// TIA Portal project "Star-Delta Motor Starter with Industrial HMI+Fault Protection" (V20)

(* hardware
DEVICE "S7-1200 station_1"  S7-1200 Station
   slot 0: "Rack_0"  S7-1200 Rack  Rack  V1.0
   slot 1: "PLC_1"  CPU 1214C DC/DC/DC  6ES7 214-1AG40-0XB0  V4.7
DEVICE "HMI_1"  KTP700 Basic PN
   slot 0: "HMI_1"  KTP700 Basic PN  6AV2 123-2GB03-0AX0  17.0.0.0
   slot 1: "HMI_RT_1"  KTP700 Basic PN  6AV2 123-2GB03-0AX0  17.0.0.0
   slot 5: "HMI_1.IE_CP_1"  PROFINET Interface  17.0.0.0
      slot 1: "PROFINET Interface_1"  PROFINET Interface
         slot 1: "Port_1"  Port
*)

// ===== PLC "PLC_1"  CPU 1214C DC/DC/DC =====

VAR_GLOBAL   // PLC tag table "Default tag table"
   "Start_PB" AT %I0.0 : Bool;
   "Stop_PB" AT %I0.1 : Bool;
   "Emergency_Stop" AT %I0.2 : Bool;
   "Thermal_Overload" AT %I0.3 : Bool;
   "Phase_Loss_Sensor" AT %I0.4 : Bool;
   "Reset_PB" AT %I0.5 : Bool;
   "Main_Contactor_K1" AT %Q0.0 : Bool;
   "Star_Contactor_K2" AT %Q0.1 : Bool;
   "Delta_Contactor_K3" AT %Q0.2 : Bool;
   "Alarm_Lamp" AT %M10.3 : Bool;
   "Motor_Run_Latch" AT %M0.0 : Bool;
   "Star_Mode" AT %M0.1 : Bool;
   "Delta_Mode" AT %M0.2 : Bool;
   "Fault_Active" AT %M0.3 : Bool;
   "HMI_Start" AT %M0.4 : Bool;
   "HMI_Stop" AT %M0.5 : Bool;
   "HMI_Reset" AT %M0.6 : Bool;
   "Transition_Done" AT %M0.7 : Bool;
   "Start_Command" AT %M1.0 : Bool;
   "Stop_Command" AT %M1.1 : Bool;
   "Star_Timer_Done" AT %M1.2 : Bool;
   "Star_Lamp" AT %M10.2 : Bool;
   "Delta_Lamp" AT %M10.1 : Bool;
   "Start_Pulse" AT %M1.3 : Bool;
END_VAR

DATA_BLOCK "DB_StarDelta"   // DB1
{ S7_Optimized_Access := 'TRUE' }
VERSION : 0.1
   VAR
      Star_timer_Preset : Time := T#5s;
      Transition_Delay : Time := T#500ms;
      Running_Hours : Real := 0.0;
      Start_Counter : Int := 0;
      Fault_Code : Int := 0;
      Motor_Status : Bool;
      Thermal_Alarm : Bool;
      Phase_Loss_Alarm : Bool;
      Star_Contactor_Fault : Bool;
      Delta_Contactor_Fault : Bool;
   END_VAR
BEGIN
END_DATA_BLOCK

// folder: System blocks/Program resources

DATA_BLOCK "Star_Timer"   // DB2
{ S7_Optimized_Access := 'TRUE' }
AUTHOR : Simatic
FAMILY : IEC
NAME : IEC_TMR
VERSION : 1.0
// stored: InstanceOfName IEC_TIMER
"IEC_TIMER"
BEGIN
END_DATA_BLOCK

DATA_BLOCK "Transition_Timer"   // DB3
{ S7_Optimized_Access := 'TRUE' }
AUTHOR : Simatic
FAMILY : IEC
NAME : IEC_TMR
VERSION : 1.0
// stored: InstanceOfName IEC_TIMER
"IEC_TIMER"
BEGIN
END_DATA_BLOCK

// folder: (top level)

ORGANIZATION_BLOCK "Main"   // OB1, LAD, ProgramCycle
TITLE = "Main Program Sweep (Cycle)"
{ S7_Optimized_Access := 'TRUE' }
VERSION : 0.1
   VAR_INPUT
      Initial_Call : Bool;   // Initial call of this OB
      Remanence : Bool;   // =True, if remanent data are available
   END_VAR
BEGIN

REGION Network 1: Start command
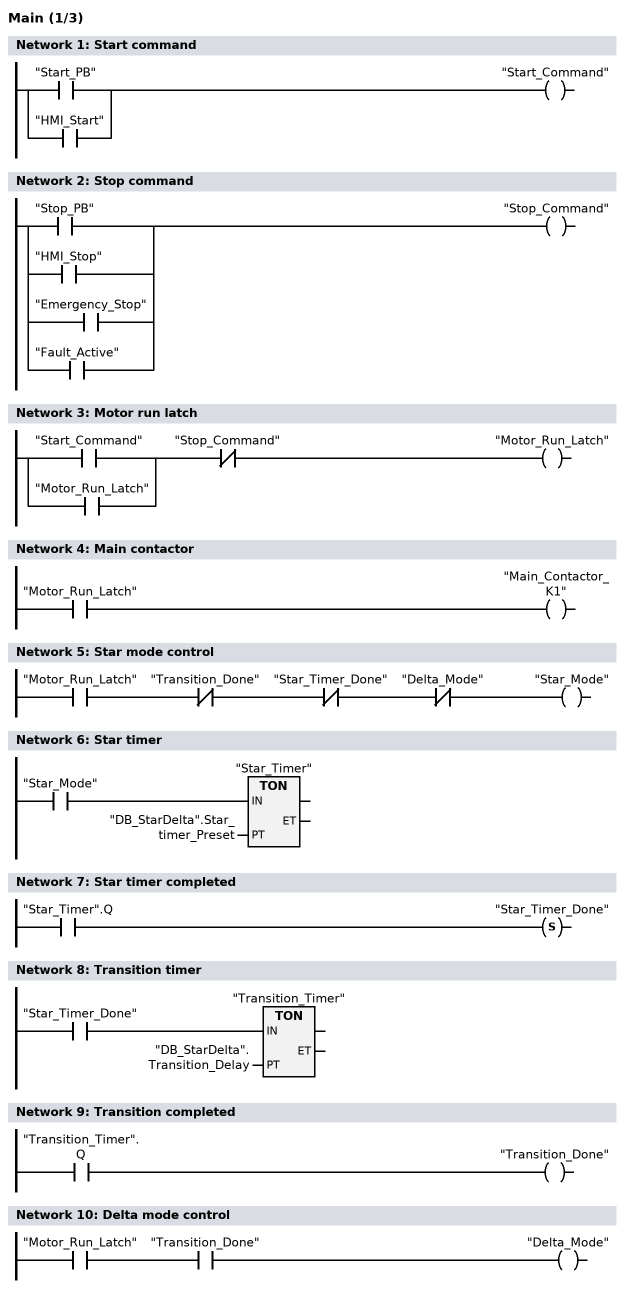
   RUNG wire#powerrail
      Contact( "Start_PB" )
      wire#w1
      Coil( "Start_Command" )
   END_RUNG
   RUNG wire#powerrail
      Contact( "HMI_Start" )
   END_RUNG wire#w1
   // the same network as SCL:
   "Start_Command" := "Start_PB" OR "HMI_Start";
END_REGION

REGION Network 2: Stop command
   RUNG wire#powerrail
      Contact( "Stop_PB" )
      wire#w1
      Coil( "Stop_Command" )
   END_RUNG
   RUNG wire#powerrail
      Contact( "HMI_Stop" )
   END_RUNG wire#w1
   RUNG wire#powerrail
      Contact( "Emergency_Stop" )
   END_RUNG wire#w1
   RUNG wire#powerrail
      Contact( "Fault_Active" )
   END_RUNG wire#w1
   // the same network as SCL:
   "Stop_Command" := "Stop_PB" OR "HMI_Stop" OR "Emergency_Stop" OR "Fault_Active";
END_REGION

REGION Network 3: Motor run latch
   RUNG wire#powerrail
      Contact( "Start_Command" )
      wire#w1
      I_Contact( "Stop_Command" )
      Coil( "Motor_Run_Latch" )
   END_RUNG
   RUNG wire#powerrail
      Contact( "Motor_Run_Latch" )
   END_RUNG wire#w1
   // the same network as SCL:
   "Motor_Run_Latch" := ("Start_Command" OR "Motor_Run_Latch") AND NOT "Stop_Command";
END_REGION

REGION Network 4: Main contactor
   RUNG wire#powerrail
      Contact( "Motor_Run_Latch" )
      Coil( "Main_Contactor_K1" )
   END_RUNG
   // the same network as SCL:
   "Main_Contactor_K1" := "Motor_Run_Latch";
END_REGION

REGION Network 5: Star mode control
   RUNG wire#powerrail
      Contact( "Motor_Run_Latch" )
      I_Contact( "Transition_Done" )
      I_Contact( "Star_Timer_Done" )
      I_Contact( "Delta_Mode" )
      Coil( "Star_Mode" )
   END_RUNG
   // the same network as SCL:
   "Star_Mode" := "Motor_Run_Latch" AND NOT "Transition_Done" AND NOT "Star_Timer_Done" AND NOT "Delta_Mode";
END_REGION

REGION Network 6: Star timer
   "Star_Timer".TON(IN := "Star_Mode", PT := "DB_StarDelta".Star_timer_Preset);
END_REGION

REGION Network 7: Star timer completed
   RUNG wire#powerrail
      Contact( "Star_Timer".Q )
      S_Coil( "Star_Timer_Done" )
   END_RUNG
   // the same network as SCL:
   IF "Star_Timer".Q THEN "Star_Timer_Done" := TRUE; END_IF;
END_REGION

REGION Network 8: Transition timer
   "Transition_Timer".TON(IN := "Star_Timer_Done", PT := "DB_StarDelta".Transition_Delay);
END_REGION

REGION Network 9: Transition completed
   RUNG wire#powerrail
      Contact( "Transition_Timer".Q )
      Coil( "Transition_Done" )
   END_RUNG
   // the same network as SCL:
   "Transition_Done" := "Transition_Timer".Q;
END_REGION

REGION Network 10: Delta mode control
   RUNG wire#powerrail
      Contact( "Motor_Run_Latch" )
      Contact( "Transition_Done" )
      Coil( "Delta_Mode" )
   END_RUNG
   // the same network as SCL:
   "Delta_Mode" := "Motor_Run_Latch" AND "Transition_Done";
END_REGION

REGION Network 11: Delta contactor
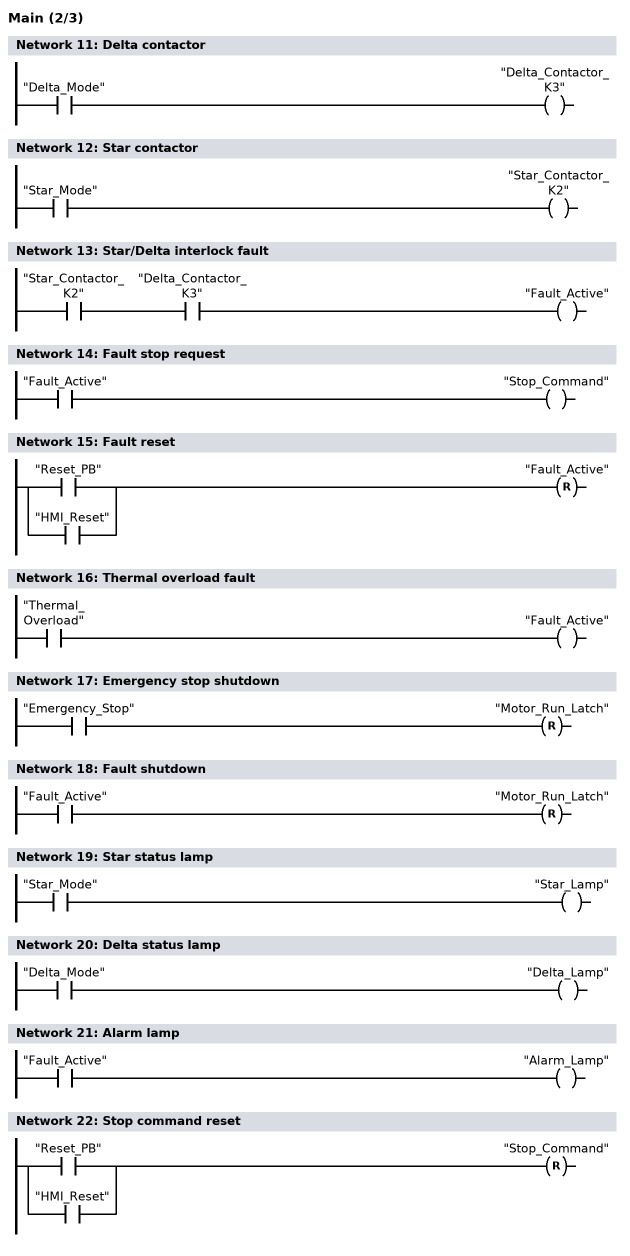
   RUNG wire#powerrail
      Contact( "Delta_Mode" )
      Coil( "Delta_Contactor_K3" )
   END_RUNG
   // the same network as SCL:
   "Delta_Contactor_K3" := "Delta_Mode";
END_REGION

REGION Network 12: Star contactor
   RUNG wire#powerrail
      Contact( "Star_Mode" )
      Coil( "Star_Contactor_K2" )
   END_RUNG
   // the same network as SCL:
   "Star_Contactor_K2" := "Star_Mode";
END_REGION

REGION Network 13: Star/Delta interlock fault
   RUNG wire#powerrail
      Contact( "Star_Contactor_K2" )
      Contact( "Delta_Contactor_K3" )
      Coil( "Fault_Active" )
   END_RUNG
   // the same network as SCL:
   "Fault_Active" := "Star_Contactor_K2" AND "Delta_Contactor_K3";
END_REGION

REGION Network 14: Fault stop request
   RUNG wire#powerrail
      Contact( "Fault_Active" )
      Coil( "Stop_Command" )
   END_RUNG
   // the same network as SCL:
   "Stop_Command" := "Fault_Active";
END_REGION

REGION Network 15: Fault reset
   RUNG wire#powerrail
      Contact( "Reset_PB" )
      wire#w1
      R_Coil( "Fault_Active" )
   END_RUNG
   RUNG wire#powerrail
      Contact( "HMI_Reset" )
   END_RUNG wire#w1
   // the same network as SCL:
   IF "Reset_PB" OR "HMI_Reset" THEN "Fault_Active" := FALSE; END_IF;
END_REGION

REGION Network 16: Thermal overload fault
   RUNG wire#powerrail
      Contact( "Thermal_Overload" )
      Coil( "Fault_Active" )
   END_RUNG
   // the same network as SCL:
   "Fault_Active" := "Thermal_Overload";
END_REGION

REGION Network 17: Emergency stop shutdown
   RUNG wire#powerrail
      Contact( "Emergency_Stop" )
      R_Coil( "Motor_Run_Latch" )
   END_RUNG
   // the same network as SCL:
   IF "Emergency_Stop" THEN "Motor_Run_Latch" := FALSE; END_IF;
END_REGION

REGION Network 18: Fault shutdown
   RUNG wire#powerrail
      Contact( "Fault_Active" )
      R_Coil( "Motor_Run_Latch" )
   END_RUNG
   // the same network as SCL:
   IF "Fault_Active" THEN "Motor_Run_Latch" := FALSE; END_IF;
END_REGION

REGION Network 19: Star status lamp
   RUNG wire#powerrail
      Contact( "Star_Mode" )
      Coil( "Star_Lamp" )
   END_RUNG
   // the same network as SCL:
   "Star_Lamp" := "Star_Mode";
END_REGION

REGION Network 20: Delta status lamp
   RUNG wire#powerrail
      Contact( "Delta_Mode" )
      Coil( "Delta_Lamp" )
   END_RUNG
   // the same network as SCL:
   "Delta_Lamp" := "Delta_Mode";
END_REGION

REGION Network 21: Alarm lamp
   RUNG wire#powerrail
      Contact( "Fault_Active" )
      Coil( "Alarm_Lamp" )
   END_RUNG
   // the same network as SCL:
   "Alarm_Lamp" := "Fault_Active";
END_REGION

REGION Network 22: Stop command reset
   RUNG wire#powerrail
      Contact( "Reset_PB" )
      wire#w1
      R_Coil( "Stop_Command" )
   END_RUNG
   RUNG wire#powerrail
      Contact( "HMI_Reset" )
   END_RUNG wire#w1
   // the same network as SCL:
   IF "Reset_PB" OR "HMI_Reset" THEN "Stop_Command" := FALSE; END_IF;
END_REGION

REGION Network 23: Transition flag reset
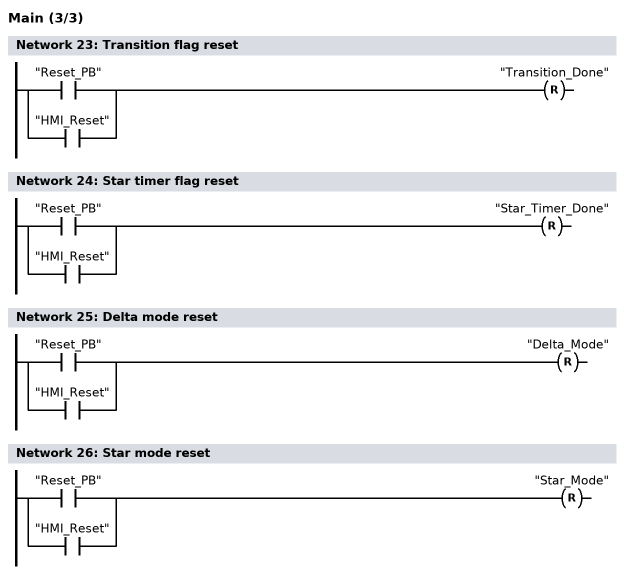
   RUNG wire#powerrail
      Contact( "Reset_PB" )
      wire#w1
      R_Coil( "Transition_Done" )
   END_RUNG
   RUNG wire#powerrail
      Contact( "HMI_Reset" )
   END_RUNG wire#w1
   // the same network as SCL:
   IF "Reset_PB" OR "HMI_Reset" THEN "Transition_Done" := FALSE; END_IF;
END_REGION

REGION Network 24: Star timer flag reset
   RUNG wire#powerrail
      Contact( "Reset_PB" )
      wire#w1
      R_Coil( "Star_Timer_Done" )
   END_RUNG
   RUNG wire#powerrail
      Contact( "HMI_Reset" )
   END_RUNG wire#w1
   // the same network as SCL:
   IF "Reset_PB" OR "HMI_Reset" THEN "Star_Timer_Done" := FALSE; END_IF;
END_REGION

REGION Network 25: Delta mode reset
   RUNG wire#powerrail
      Contact( "Reset_PB" )
      wire#w1
      R_Coil( "Delta_Mode" )
   END_RUNG
   RUNG wire#powerrail
      Contact( "HMI_Reset" )
   END_RUNG wire#w1
   // the same network as SCL:
   IF "Reset_PB" OR "HMI_Reset" THEN "Delta_Mode" := FALSE; END_IF;
END_REGION

REGION Network 26: Star mode reset
   RUNG wire#powerrail
      Contact( "Reset_PB" )
      wire#w1
      R_Coil( "Star_Mode" )
   END_RUNG
   RUNG wire#powerrail
      Contact( "HMI_Reset" )
   END_RUNG wire#w1
   // the same network as SCL:
   IF "Reset_PB" OR "HMI_Reset" THEN "Star_Mode" := FALSE; END_IF;
END_REGION
END_ORGANIZATION_BLOCK

(* ===== HMI "HMI_RT_1" =====
system functions are stored by id; their names below are inferred from use
connection "HMI_Connection_1": ETHERNET, SMART_S7_1200_OMS

HMI tags "Default tag table"
   "Tag_ScreenNumber" : UInt, internal
   "Fault_Active" : Bool = PLC Fault_Active AT %M0.3, 1 s
   "Main_Contactor_K1" : Bool = PLC Main_Contactor_K1 AT %Q0.0, 1 s
   "HMI_Start" : Bool = PLC HMI_Start AT %M0.4, 1 s
   "HMI_Stop" : Bool = PLC HMI_Stop AT %M0.5, 1 s
   "HMI_Reset" : Bool = PLC HMI_Reset AT %M0.6, 1 s
   "Emergency_Stop" : Bool = PLC Emergency_Stop AT %I0.2, 1 s
   "Delta_Mode" : Bool = PLC Delta_Mode AT %M0.2, 1 s
   "Star_Contactor_K2" : Bool = PLC Star_Contactor_K2 AT %Q0.1, 1 s
   "Delta_Contactor_K3" : Bool = PLC Delta_Contactor_K3 AT %Q0.2, 1 s

text list "ON": 0 'OFF'; 1 'ON'

Template "Template_1" 800x480
   Button "Exit" at 714,429 size 71x50; TextOff 'Exit'; PictureOff "ExitRuntime_KTP700_Basic_PN_TR"; PictureOn "ExitRuntime_KTP700_Basic_PN_TR"
      on Release: StopRuntime(0)
   Button "Template_Button" at 614,429 size 71x50; TextOff 'Text'
   Button "Template_Button_1" at 514,429 size 71x50; TextOff 'Text'
   Button "Template_Button_2" at 414,429 size 71x50; TextOff 'Text'
   Button "Template_Button_3" at 314,429 size 71x50; TextOff 'Text'
   Button "Template_Button_4" at 214,429 size 71x50; TextOff 'Text'
   Button "Template_Button_5" at 114,429 size 71x50; TextOff 'Text'
   Button "Start screen" at 14,429 size 71x50; TextOff 'Start screen'; PictureOff "NavigateHome_KTP700_Basic_PN_TR"; PictureOn "NavigateHome_KTP700_Basic_PN_TR"
      on Release: ActivateScreen("Main Overview", 0)
   SymbolicIOField "Symbolic_IO_Field_Screen" at 93,9 size 600x33; TextOff '0'; TextOn '1'; TextList "TextList_ScreenNames"
      ProcessValue <- "Tag_ScreenNumber"
      on Change: ActivateScreenByNumber("Tag_ScreenNumber", 0)
   DateTimeField "HmiScreenItemData" at 695,25 size 105x25
   DateTimeField "HmiScreenItemData_1" at 695,0 size 105x25
   GraphicView "Logo" at 0,0 size 91x51; Picture "Logo of HMI_1"

screen "Main Overview" 800x480, template "Template_1"
   on GenerateScreen: SetTag("Tag_ScreenNumber", 1)
   GraphicView "Graphic view_1" at 0,0 size 800x479; Picture "ChatGPT Image 25 Ιουν 2026, 09_10_57 μ.μ."
   TextField "Text field_1" at 240,213 size 80x36; Text 'MAIN CONTACTOR'
   Button "Button_1" at 0,431 size 195x48; TextOff 'MAIN OVERVIEW'
   Button "Button_2" at 195,431 size 195x48; TextOff 'CONTROL'
   Button "Button_3" at 389,431 size 191x48; TextOff 'ALARMS'
   Button "Button_4" at 580,431 size 219x48; TextOff 'DIAGNOSTICS'
   Button "Button_5" at 77,360 size 195x48; TextOff 'START'
      on Press: function_b14e0dd5("HMI_Start", 0)
   Button "Button_6" at 307,359 size 195x48; TextOff 'STOP'
      on Press: function_b14e0dd5("HMI_Stop", 0)
   Button "Button_7" at 532,360 size 195x48; TextOff 'RESET'
      on Press: function_b14e0dd5("HMI_Reset", 0)
   GraphicView "Graphic view_2" at 235,247 size 93x74; Picture "κ1_1"
   GraphicView "Graphic view_3" at 336,248 size 82x74; Picture "κ1_1"
   GraphicView "Graphic view_4" at 430,248 size 82x74; Picture "κ1_1"
   TextField "Text field_2" at 55,102 size 125x22; Text 'MOTOR STATUS'
   TextField "Text field_3" at 55,163 size 133x22; Text 'STARTING MODE'
   TextField "Text field_4" at 55,222 size 121x22; Text 'ALARM STATUS'
   TextField "Text field_5" at 55,282 size 124x22; Text 'E-STOP STATUS'
   GraphicView "Graphic view_5" at 603,437 size 36x30; Picture "Graphic_1"
   GraphicView "Graphic view_6" at 415,439 size 36x30; Picture "Graphic_2"
   GraphicView "Graphic view_7" at 19,229 size 36x30; Picture "Graphic_2"
      Appearance <- "Fault_Active"
   GraphicView "Graphic view_8" at -1,439 size 36x30; Picture "Graphic_3"
   GraphicView "Graphic view_10" at 215,439 size 36x30; Picture "Graphic_5"
   GraphicView "Graphic view_11" at 257,34 size 232x156; Picture "μοτορ"
   TextField "Text field_6" at 265,189 size 21x20; Text 'K1'
   TextField "Text field_7" at 336,213 size 80x36; Text 'STAR CONTACTOR'
   TextField "Text field_8" at 361,191 size 21x20; Text 'K2'
   TextField "Text field_9" at 430,213 size 80x36; Text 'DELTA CONTACTOR'
   TextField "Text field_10" at 456,191 size 21x20; Text 'K3'
   TextField "Text field_11" at 254,2 size 237x22; Text 'STAR-DELTA MOTOR STARTER'
   GraphicView "Graphic view_12" at 19,171 size 36x30; Picture "Graphic_6"
      Appearance <- "Delta_Mode"
   GraphicView "Graphic view_9" at 18,294 size 36x30; Picture "Graphic_7"
   SymbolicIOField "Symbolic I/O field_1" at 254,321 size 52x23; TextOff '0'; TextOn '1'; TextList "ON"
      ProcessValue <- "Main_Contactor_K1"
      Appearance <- "Main_Contactor_K1"
   SymbolicIOField "Symbolic I/O field_2" at 348,322 size 52x23; TextOff '0'; TextOn '1'; TextList "ON"
      ProcessValue <- "Star_Contactor_K2"
      Appearance <- "Star_Contactor_K2"
   SymbolicIOField "Symbolic I/O field_3" at 445,322 size 52x23; TextOff '0'; TextOn '1'; TextList "ON"
      ProcessValue <- "Delta_Contactor_K3"
      Appearance <- "Delta_Contactor_K3"
   SymbolicIOField "Symbolic I/O field_4" at 58,304 size 52x28; TextOff '0'; TextOn '1'; TextList "ON"
      ProcessValue <- "Emergency_Stop"
   TextField "Text field_12" at 55,244 size 29x22; Text 'NO'
      Visibility <- "Fault_Active"
   TextField "Text field_13" at 83,244 size 53x22; Text 'FAULT'
      Appearance <- "Fault_Active"
   TextField "Text field_14" at 585,106 size 34x37; Text '1)'
   TextField "Text field_15" at 616,102 size 112x46; Text 'MAIN+STAR K1+K2 ON'
   GraphicView "Graphic view_13" at 646,154 size 36x30; Picture "Graphic_8"
   GraphicView "Graphic view_14" at 646,237 size 36x30; Picture "Graphic_8"
   TextField "Text field_16" at 586,191 size 34x37; Text '2)'
   TextField "Text field_17" at 621,189 size 120x46; Text 'TRANSITION DELAY(T1)'
   TextField "Text field_18" at 621,276 size 122x46; Text 'MAIN+DELTA K1+K3 ON'
   TextField "Text field_19" at 585,278 size 34x37; Text '3)'
   TextField "Text field_20" at 580,61 size 170x22; Text 'STARTING SEQUENCE'

screen "Control" 800x480, template "Template_1"
   on GenerateScreen: SetTag("Tag_ScreenNumber", 2)
   TextField "HmiScreenItemData" at 80,225 size 640x25; Text 'Control'
   Button "Back" at 1,52 size 159x47; TextOff 'Back'
      on Release: ActivateScreen("Main Overview", 0)

screen "Alarm Page" 800x480, template "Template_1"
   on GenerateScreen: SetTag("Tag_ScreenNumber", 3)
   TextField "HmiScreenItemData" at 80,225 size 640x25; Text 'Alarm Page'
   Button "Back" at 1,52 size 159x47; TextOff 'Back'
      on Release: ActivateScreen("Main Overview", 0)

screen "Diagnostics" 800x480, template "Template_1"
   on GenerateScreen: SetTag("Tag_ScreenNumber", 4)
   TextField "HmiScreenItemData" at 80,225 size 640x25; Text 'Diagnostics'
   Button "Back" at 1,52 size 159x47; TextOff 'Back'
      on Release: ActivateScreen("Main Overview", 0)
*)